(* Logix 5000 project; controller MV vendor 1 type 14 code 217 rev 31.11; software revision 31.00; part 43 of 53 *)
(* tags used below, declared in another part *)
   Always_Off : BOOL;
   CWD : CHECKWORD_FLAGS;
   Enable_TimeString : BOOL;
   MC_N100 : INT[255];   // C1_PLC Channel 1 PLC data
   MC_N120 : INT[255];   // C2 PLC Channel 2 PLC data
   MV_BM01_AV01 : PlantItem;   // BM01_AV01
   MV_BM01_AV01_CIP : BOOL;
   MV_BM01_AV01_MV20 : BOOL;
   MV_BM01_ZS04 : PlantItem;   // BM01ZS04
   MV_BM01_ZS05 : PlantItem;   // BM01ZS05
   MV_DAL01_AV01_MV20 : BOOL;
   MV_Data_To_TF : DINT[30];
   MV_Enable_MV20_NewPressureControl : BOOL;
   MV_FP01_ZS01 : PlantItem;   // FP01ZS01
   MV_FP01_ZS02 : PlantItem;   // FP01ZS02
   MV_GasAvailable : BOOL;
   MV_MV20_AV01 : PlantItem;   // MV20_AV01
   MV_MV20_CIP : BOOL;
   MV_MV20_CO2 : BOOL;
   MV_MV20_CO2_ON_PreStorage : BOOL;
   MV_MV20_CO2_ON_Storage : BOOL;
   MV_MV20_ControlOpenVent : BOOL;
   MV_MV20_Filling_Pulse : BOOL;
   MV_MV20_Filling_PulseLevel : REAL;
   MV_MV20_LTX07_TrueLevel : REAL;
   MV_MV20_ProxiesOK : BOOL;
   MV_MV20_PTX01_AI : PlantItem;   // MV20_PTX01
   MV_MV20_TP_CaskDepressure : BOOL;
   MV_MV20_TP_CaskEmptying : BOOL;
   MV_MV20_TP_CaskFilling : BOOL;
   MV_MV20_TP_CaskPreEmptyPressure : BOOL;
   MV_MV20_TP_CaskPrePressure : BOOL;
   MV_MV20_TP_CaskPressureDelay : BOOL;
   MV_MV20_TP_CaskPurgeFromTop : BOOL;
   MV_MV20_TP_CaskReadyToFill : BOOL;
   MV_MV20_TP_CaskStorage : BOOL;
   MV_MV20_TP_CO2_Debounce_Timer : TIMER;
   MV_MV20_TP_CO2_Debounce_Timer_1 : TIMER;
   MV_MV20_TP_CO2_HSL_Pressure : REAL;
   MV_MV20_TP_CO2_HSL_Storage : REAL;
   MV_MV20_TP_CO2_HSL_Timer : TIMER;
   MV_MV20_TP_CO2_LSL_pressure_1 : REAL;
   MV_MV20_TP_CO2_LSL_storage : REAL;
   MV_MV20_TP_CO2_LSL_Timer : TIMER;
   MV_MV20_TP_Command : DINT;
   MV_MV20_TP_DAL_Chase_Cask : BOOL;
   MV_MV20_TP_DAL_Chase_KB : BOOL;
   MV_MV20_TP_DAL_Chase_Time : TIMER;
   MV_MV20_TP_Dirty : BOOL;
   MV_MV20_TP_Emptying_Level_Setpoint : REAL;
   MV_MV20_TP_Error_String : STRING;
   MV_MV20_TP_Faulted : BOOL;
   MV_MV20_TP_Fill_Pulse_OFF_Timer : TIMER;
   MV_MV20_TP_Fill_Pulse_ON_Timer : TIMER;
   MV_MV20_TP_Held : BOOL;
   MV_MV20_TP_Idle : BOOL;
   MV_MV20_TP_Initial_DAL_Chase_Cask : BOOL;
   MV_MV20_TP_Initial_DAL_Chase_KB : BOOL;
   MV_MV20_TP_KBEmptying : BOOL;
   MV_MV20_TP_KBFilling : BOOL;
   MV_MV20_TP_KBFillingBuildPressure : BOOL;
   MV_MV20_TP_KBPreEmptyPressure : BOOL;
   MV_MV20_TP_KBPrePressurise : BOOL;
   MV_MV20_TP_KBStorage : BOOL;
   MV_MV20_TP_LowerLimit : REAL;
   MV_MV20_TP_ONS_1 : BOOL;
   MV_MV20_TP_Prompt : DINT;
   MV_MV20_TP_Proxy_Delay_Made : TIMER;
   MV_MV20_TP_Proxy_Delay_NOT_MADE : TIMER;
   MV_MV20_TP_Pulse : BOOL;
   MV_MV20_TP_ReadyToFillKB : BOOL;
   MV_MV20_TP_ReadyToFillKB_M : BOOL;
   MV_MV20_TP_Running : BOOL;
   MV_MV20_TP_Setpoint : REAL;
   MV_MV20_TP_Status : DINT;   // 0 = Idle, 1 = Running, 2 = Held, 3 = Faulted
   MV_MV20_TP_Step : DINT;
   MV_MV20_TP_Steptime : DINT;
   MV_MV20_TP_Steptime_String : STRING;
   MV_MV20_TP_SteptimeRunning : DINT;
   MV_MV20_TP_TimeLeft : DINT;
   MV_MV20_TP_TimeLeft_msec : DINT;
   MV_MV20_TP_TimeLeftStr : STRING;
   MV_MV20_TP_UpperLimit : REAL;
   MV_MV20_TP_Vent : BOOL;
   MV_MV20_TPLastStep : DINT;
   MV_MV20_Transfer_StartLevel : REAL;
   MV_MV20_Transferred_Level : REAL;
   MV_MV21_TP_Status : DINT;   // 0 = Idle, 1 = Running, 2 = Held, 3 = Faulted
   MV_N136 : INT[50];   // MV 20, CURRENT FV DATA
   MV_TP_CaskEmptyingPressure : REAL;
   MV_TP_CaskFillingPressure : REAL;
   MV_TP_CaskPrefillPressure : REAL;
   MV_TP_CaskStoragePressure : REAL;
   MV_TP_CaskStoragePressureDelay : DINT;
   MV_TP_CaskStoragePressureDelay_Secs : DINT;
   MV_TP_CaskStoragePressureLevel : REAL;
   MV_TP_Deadband : REAL;
   MV_TP_Emptying_Volume_Setpoint : REAL;
   MV_TP_HighLevelDeadband : REAL;
   MV_TP_KBFillingPressure : REAL;
   MV_TP_KBStoragePressure : REAL;
   MV_TP_LowLevelDeadbandThreshold : REAL;
   MV_TP_VentPressure : REAL;
   One_Second_1_scan : BOOL;
(* MV_Common, continued *)

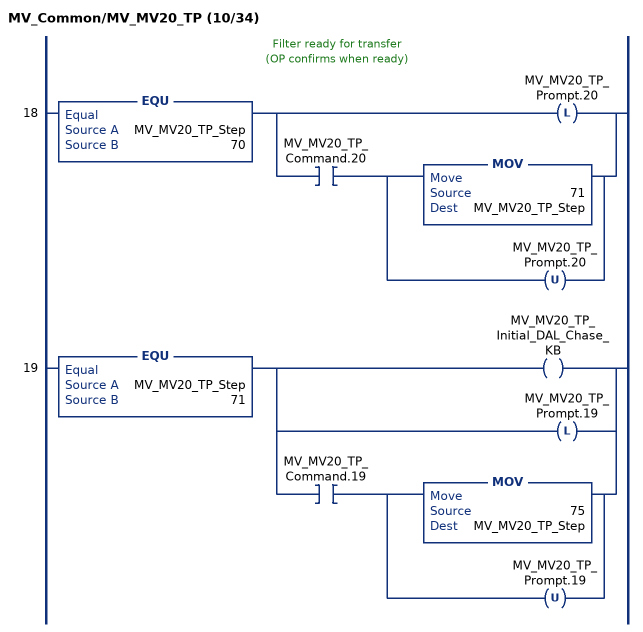
   // Filter ready for transfer
   // (OP confirms when ready)
   18: EQU(MV_MV20_TP_Step,70)[OTL(MV_MV20_TP_Prompt.20) ,XIC(MV_MV20_TP_Command.20) [MOV(71,MV_MV20_TP_Step) ,OTU(MV_MV20_TP_Prompt.20) ] ];
   19: EQU(MV_MV20_TP_Step,71)[OTE(MV_MV20_TP_Initial_DAL_Chase_KB) ,OTL(MV_MV20_TP_Prompt.19) ,XIC(MV_MV20_TP_Command.19) [MOV(75,MV_MV20_TP_Step) ,OTU(MV_MV20_TP_Prompt.19) ] ];
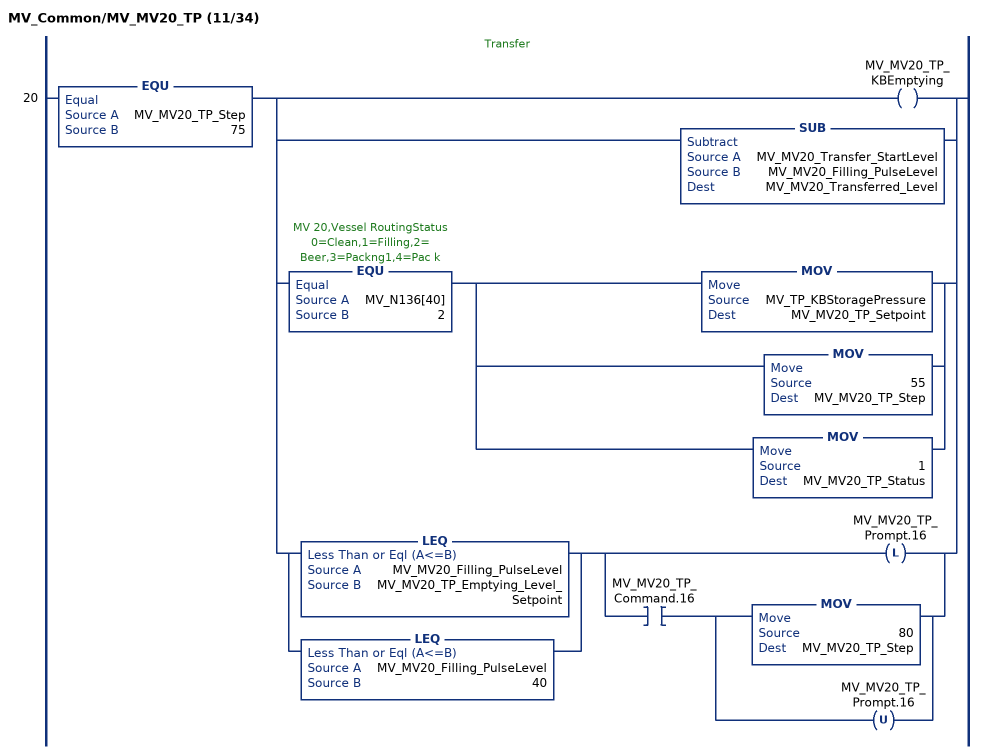
   // Transfer
   20: EQU(MV_MV20_TP_Step,75)[OTE(MV_MV20_TP_KBEmptying) ,SUB(MV_MV20_Transfer_StartLevel,MV_MV20_Filling_PulseLevel,MV_MV20_Transferred_Level) ,EQU(MV_N136[40],2) [MOV(MV_TP_KBStoragePressure,MV_MV20_TP_Setpoint) ,MOV(55,MV_MV20_TP_Step) ,MOV(1,MV_MV20_TP_Status) ] ,[LEQ(MV_MV20_Filling_PulseLevel,MV_MV20_TP_Emptying_Level_Setpoint) ,LEQ(MV_MV20_Filling_PulseLevel,40) ] [OTL(MV_MV20_TP_Prompt.16) ,XIC(MV_MV20_TP_Command.16) [MOV(80,MV_MV20_TP_Step) ,OTU(MV_MV20_TP_Prompt.16) ] ] ];
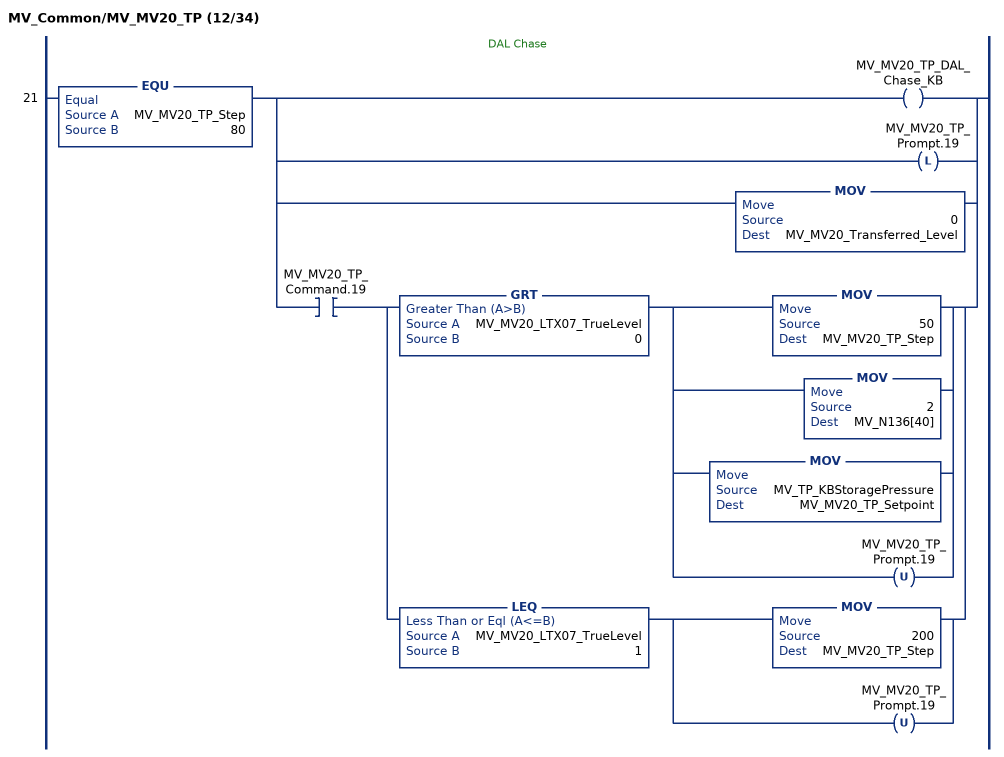
   // DAL Chase
   21: EQU(MV_MV20_TP_Step,80)[OTE(MV_MV20_TP_DAL_Chase_KB) ,OTL(MV_MV20_TP_Prompt.19) ,MOV(0,MV_MV20_Transferred_Level) ,XIC(MV_MV20_TP_Command.19) [GRT(MV_MV20_LTX07_TrueLevel,0) [MOV(50,MV_MV20_TP_Step) ,MOV(2,MV_N136[40]) ,MOV(MV_TP_KBStoragePressure,MV_MV20_TP_Setpoint) ,OTU(MV_MV20_TP_Prompt.19) ] ,LEQ(MV_MV20_LTX07_TrueLevel,1) [MOV(200,MV_MV20_TP_Step) ,OTU(MV_MV20_TP_Prompt.19) ] ] ];
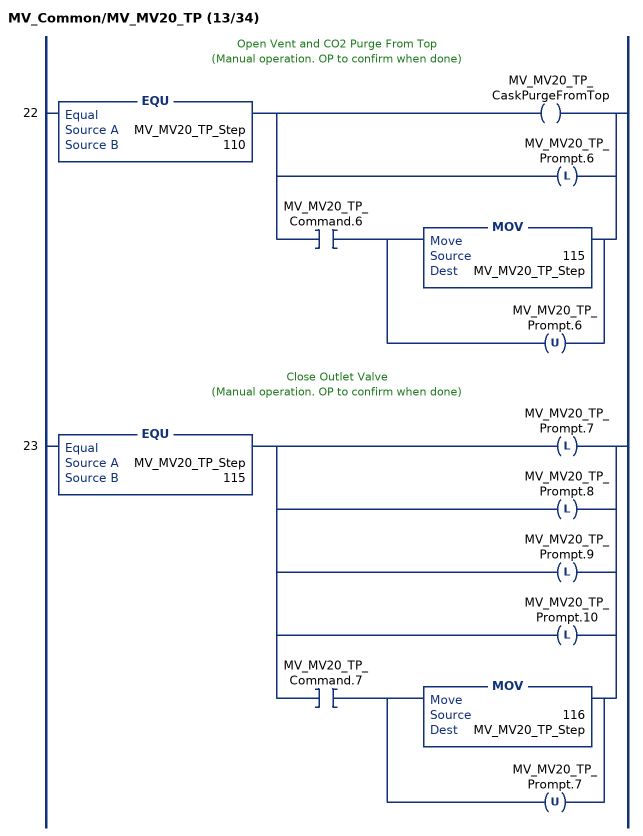
   // Open Vent and CO2 Purge From Top
   // (Manual operation. OP to confirm when done)
   22: EQU(MV_MV20_TP_Step,110)[OTE(MV_MV20_TP_CaskPurgeFromTop) ,OTL(MV_MV20_TP_Prompt.6) ,XIC(MV_MV20_TP_Command.6) [MOV(115,MV_MV20_TP_Step) ,OTU(MV_MV20_TP_Prompt.6) ] ];
   // Close Outlet Valve
   // (Manual operation. OP to confirm when done)
   23: EQU(MV_MV20_TP_Step,115)[OTL(MV_MV20_TP_Prompt.7) ,OTL(MV_MV20_TP_Prompt.8) ,OTL(MV_MV20_TP_Prompt.9) ,OTL(MV_MV20_TP_Prompt.10) ,XIC(MV_MV20_TP_Command.7) [MOV(116,MV_MV20_TP_Step) ,OTU(MV_MV20_TP_Prompt.7) ] ];
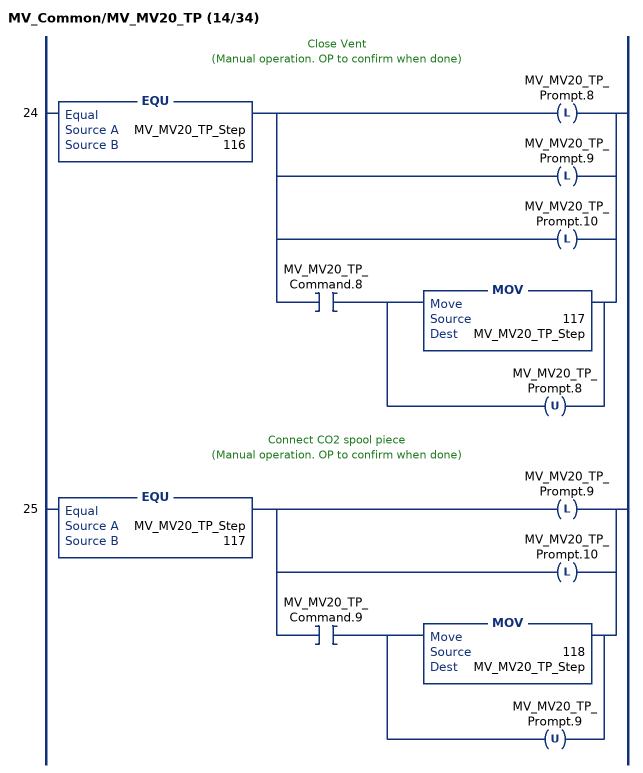
   // Close Vent
   // (Manual operation. OP to confirm when done)
   24: EQU(MV_MV20_TP_Step,116)[OTL(MV_MV20_TP_Prompt.8) ,OTL(MV_MV20_TP_Prompt.9) ,OTL(MV_MV20_TP_Prompt.10) ,XIC(MV_MV20_TP_Command.8) [MOV(117,MV_MV20_TP_Step) ,OTU(MV_MV20_TP_Prompt.8) ] ];
   // Connect CO2 spool piece
   // (Manual operation. OP to confirm when done)
   25: EQU(MV_MV20_TP_Step,117)[OTL(MV_MV20_TP_Prompt.9) ,OTL(MV_MV20_TP_Prompt.10) ,XIC(MV_MV20_TP_Command.9) [MOV(118,MV_MV20_TP_Step) ,OTU(MV_MV20_TP_Prompt.9) ] ];
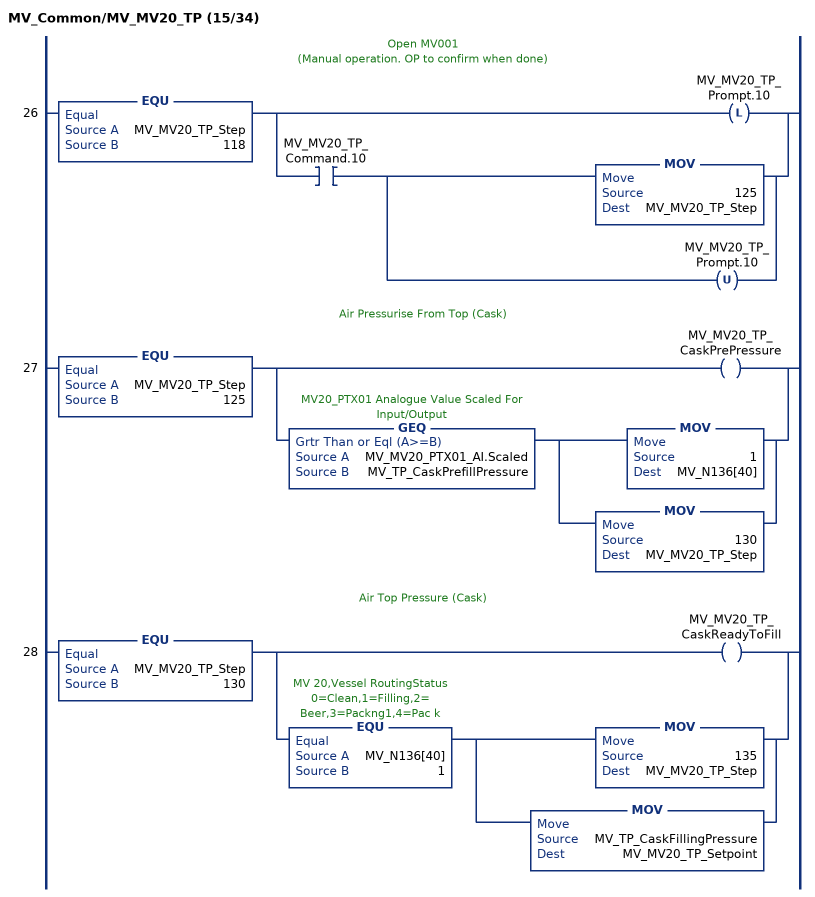
   // Open MV001
   // (Manual operation. OP to confirm when done)
   26: EQU(MV_MV20_TP_Step,118)[OTL(MV_MV20_TP_Prompt.10) ,XIC(MV_MV20_TP_Command.10) [MOV(125,MV_MV20_TP_Step) ,OTU(MV_MV20_TP_Prompt.10) ] ];
   // Air Pressurise From Top (Cask)
   27: EQU(MV_MV20_TP_Step,125)[OTE(MV_MV20_TP_CaskPrePressure) ,GEQ(MV_MV20_PTX01_AI.Scaled,MV_TP_CaskPrefillPressure) [MOV(1,MV_N136[40]) ,MOV(130,MV_MV20_TP_Step) ] ];
   // Air Top Pressure (Cask)
   28: EQU(MV_MV20_TP_Step,130)[OTE(MV_MV20_TP_CaskReadyToFill) ,EQU(MV_N136[40],1) [MOV(135,MV_MV20_TP_Step) ,MOV(MV_TP_CaskFillingPressure,MV_MV20_TP_Setpoint) ] ];
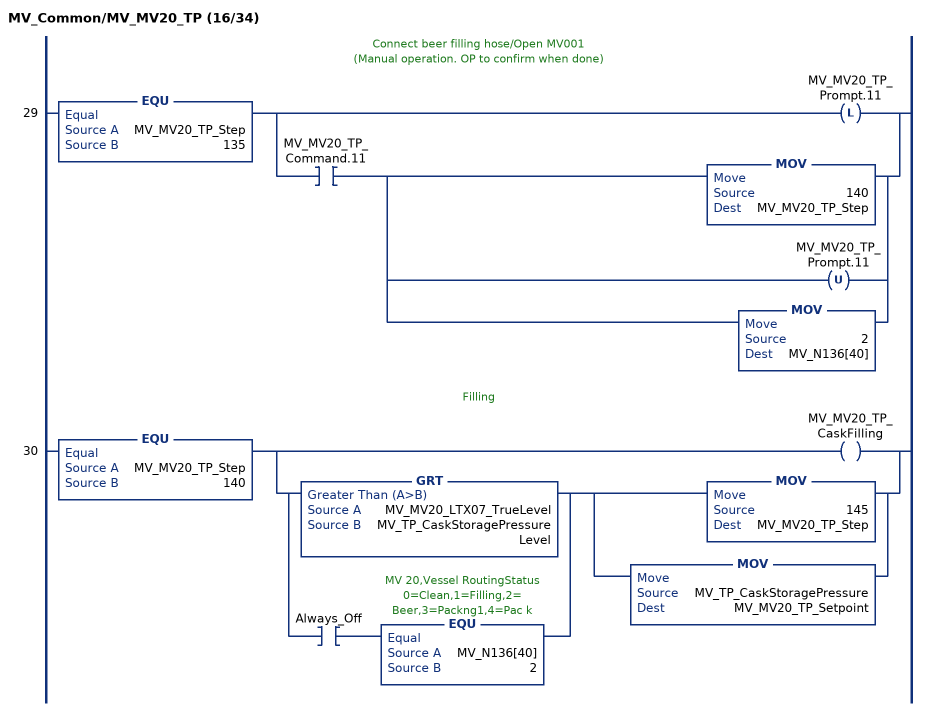
   // Connect beer filling hose/Open MV001
   // (Manual operation. OP to confirm when done)
   29: EQU(MV_MV20_TP_Step,135)[OTL(MV_MV20_TP_Prompt.11) ,XIC(MV_MV20_TP_Command.11) [MOV(140,MV_MV20_TP_Step) ,OTU(MV_MV20_TP_Prompt.11) ,MOV(2,MV_N136[40]) ] ];
   // Filling
   30: EQU(MV_MV20_TP_Step,140)[OTE(MV_MV20_TP_CaskFilling) ,[GRT(MV_MV20_LTX07_TrueLevel,MV_TP_CaskStoragePressureLevel) ,XIC(Always_Off) EQU(MV_N136[40],2) ] [MOV(145,MV_MV20_TP_Step) ,MOV(MV_TP_CaskStoragePressure,MV_MV20_TP_Setpoint) ] ];
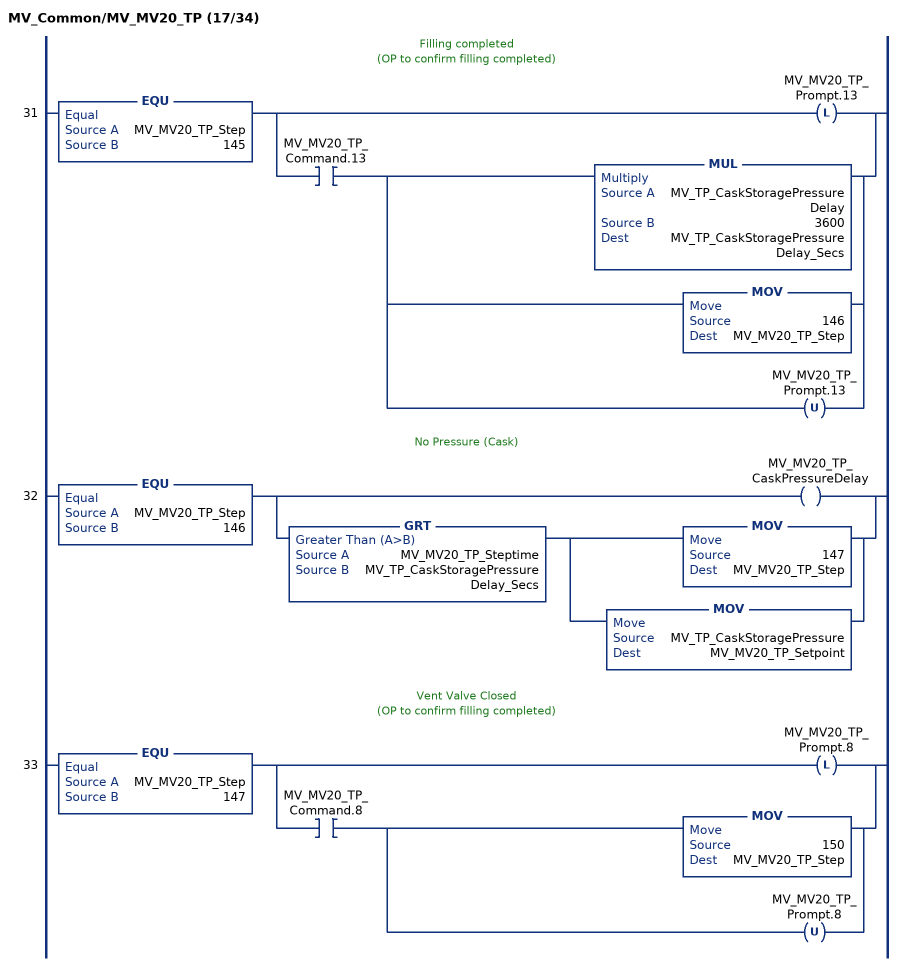
   // Filling completed
   // (OP to confirm filling completed)
   31: EQU(MV_MV20_TP_Step,145)[OTL(MV_MV20_TP_Prompt.13) ,XIC(MV_MV20_TP_Command.13) [MUL(MV_TP_CaskStoragePressureDelay,3600,MV_TP_CaskStoragePressureDelay_Secs) ,MOV(146,MV_MV20_TP_Step) ,OTU(MV_MV20_TP_Prompt.13) ] ];
   // No Pressure (Cask)
   32: EQU(MV_MV20_TP_Step,146)[OTE(MV_MV20_TP_CaskPressureDelay) ,GRT(MV_MV20_TP_Steptime,MV_TP_CaskStoragePressureDelay_Secs) [MOV(147,MV_MV20_TP_Step) ,MOV(MV_TP_CaskStoragePressure,MV_MV20_TP_Setpoint) ] ];
   // Vent Valve Closed
   // (OP to confirm filling completed)
   33: EQU(MV_MV20_TP_Step,147)[OTL(MV_MV20_TP_Prompt.8) ,XIC(MV_MV20_TP_Command.8) [MOV(150,MV_MV20_TP_Step) ,OTU(MV_MV20_TP_Prompt.8) ] ];
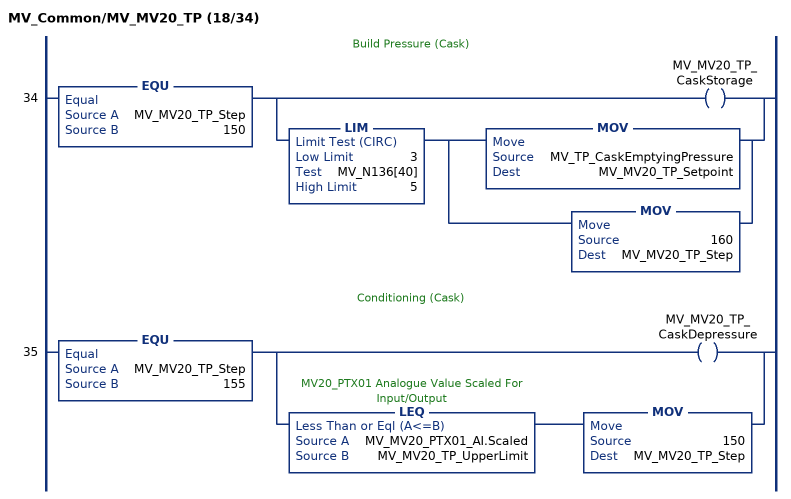
   // Build Pressure (Cask)
   34: EQU(MV_MV20_TP_Step,150)[OTE(MV_MV20_TP_CaskStorage) ,LIM(3,MV_N136[40],5) [MOV(MV_TP_CaskEmptyingPressure,MV_MV20_TP_Setpoint) ,MOV(160,MV_MV20_TP_Step) ] ];
   // Conditioning (Cask)
   35: EQU(MV_MV20_TP_Step,155)[OTE(MV_MV20_TP_CaskDepressure) ,LEQ(MV_MV20_PTX01_AI.Scaled,MV_MV20_TP_UpperLimit) MOV(150,MV_MV20_TP_Step) ];
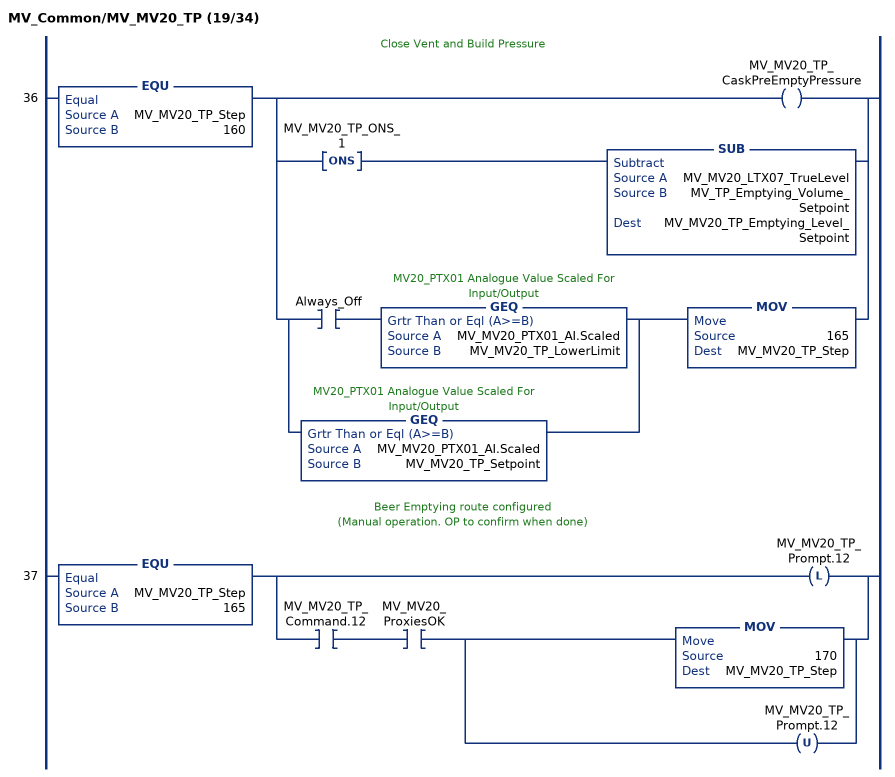
   // Close Vent and Build Pressure
   36: EQU(MV_MV20_TP_Step,160)[OTE(MV_MV20_TP_CaskPreEmptyPressure) ,ONS(MV_MV20_TP_ONS_1) SUB(MV_MV20_LTX07_TrueLevel,MV_TP_Emptying_Volume_Setpoint,MV_MV20_TP_Emptying_Level_Setpoint) ,[XIC(Always_Off) GEQ(MV_MV20_PTX01_AI.Scaled,MV_MV20_TP_LowerLimit) ,GEQ(MV_MV20_PTX01_AI.Scaled,MV_MV20_TP_Setpoint) ] MOV(165,MV_MV20_TP_Step) ];
   // Beer Emptying route configured
   // (Manual operation. OP to confirm when done)
   37: EQU(MV_MV20_TP_Step,165)[OTL(MV_MV20_TP_Prompt.12) ,XIC(MV_MV20_TP_Command.12) XIC(MV_MV20_ProxiesOK) [MOV(170,MV_MV20_TP_Step) ,OTU(MV_MV20_TP_Prompt.12) ] ];
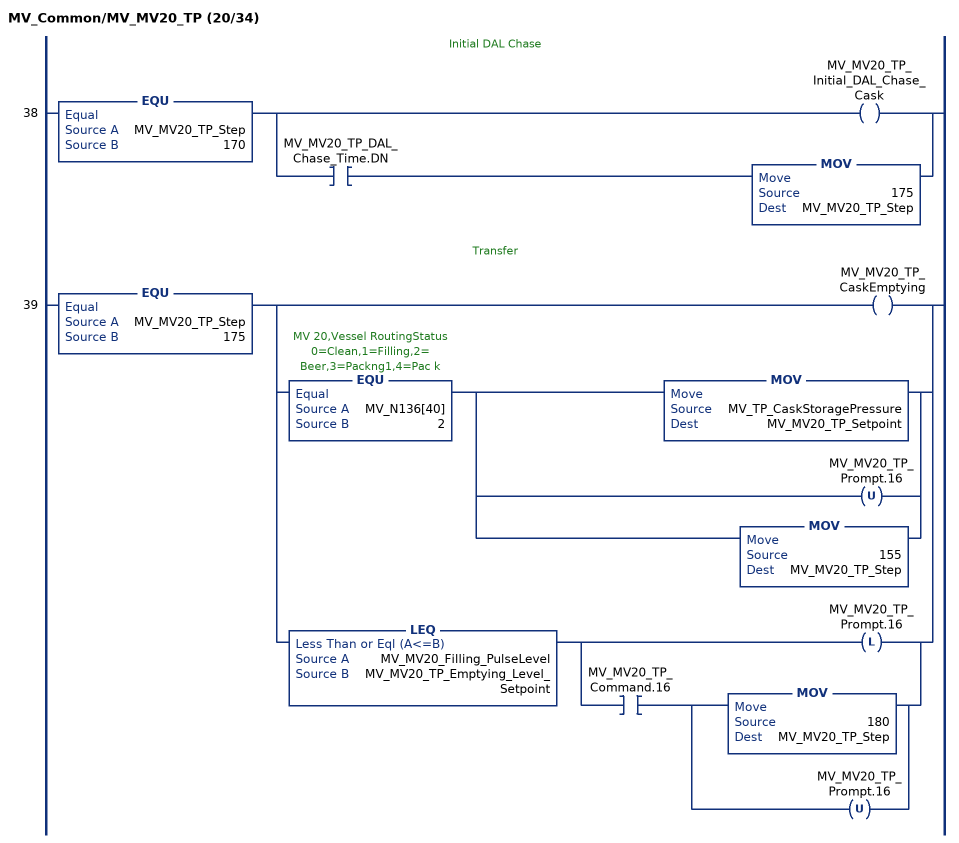
   // Initial DAL Chase
   38: EQU(MV_MV20_TP_Step,170)[OTE(MV_MV20_TP_Initial_DAL_Chase_Cask) ,XIC(MV_MV20_TP_DAL_Chase_Time.DN) MOV(175,MV_MV20_TP_Step) ];
   // Transfer
   39: EQU(MV_MV20_TP_Step,175)[OTE(MV_MV20_TP_CaskEmptying) ,EQU(MV_N136[40],2) [MOV(MV_TP_CaskStoragePressure,MV_MV20_TP_Setpoint) ,OTU(MV_MV20_TP_Prompt.16) ,MOV(155,MV_MV20_TP_Step) ] ,LEQ(MV_MV20_Filling_PulseLevel,MV_MV20_TP_Emptying_Level_Setpoint) [OTL(MV_MV20_TP_Prompt.16) ,XIC(MV_MV20_TP_Command.16) [MOV(180,MV_MV20_TP_Step) ,OTU(MV_MV20_TP_Prompt.16) ] ] ];